   
   // Copy Cap from Main line to popup
   Sbr_INO_tConvoy_SL.rgtCap[Sbr_IN_dCapIndex].dColor := Sbr_INO_tConvoyCap_ZC.rgtCap[0].dColor;
   Sbr_INO_tConvoy_SL.rgtCap[Sbr_IN_dCapIndex].dConvTotLength_cmm := Sbr_INO_tConvoyCap_ZC.rgtCap[0].dConvTotLength_cmm;
   Sbr_INO_tConvoy_SL.rgtCap[Sbr_IN_dCapIndex].dFormat := Sbr_INO_tConvoyCap_ZC.rgtCap[0].dFormat;
   Sbr_INO_tConvoy_SL.rgtCap[Sbr_IN_dCapIndex].dGap_cmm := Sbr_INO_tConvoyCap_ZC.rgtCap[0].dGap_cmm;
   Sbr_INO_tConvoy_SL.rgtCap[Sbr_IN_dCapIndex].dID := Sbr_INO_tConvoyCap_ZC.rgtCap[0].dID;
   Sbr_INO_tConvoy_SL.rgtCap[Sbr_IN_dCapIndex].dIndex := Sbr_INO_tConvoyCap_ZC.rgtCap[0].dIndex;
   Sbr_INO_tConvoy_SL.rgtCap[Sbr_IN_dCapIndex].dLength_cmm := Sbr_INO_tConvoyCap_ZC.rgtCap[0].dLength_cmm;
   Sbr_INO_tConvoy_SL.rgtCap[Sbr_IN_dCapIndex].dMaxCapInConv := Sbr_INO_tConvoyCap_ZC.rgtCap[0].dMaxCapInConv;
   Sbr_INO_tConvoy_SL.rgtCap[Sbr_IN_dCapIndex].dNumLites := Sbr_INO_tConvoyCap_ZC.rgtCap[0].dNumLites;
   Sbr_INO_tConvoy_SL.rgtCap[Sbr_IN_dCapIndex].dProductionID := Sbr_INO_tConvoyCap_ZC.rgtCap[0].dProductionID;
   Sbr_INO_tConvoy_SL.rgtCap[Sbr_IN_dCapIndex].dReqGapForConv_cmm := Sbr_INO_tConvoyCap_ZC.rgtCap[0].dReqGapForConv_cmm;
   Sbr_INO_tConvoy_SL.rgtCap[Sbr_IN_dCapIndex].dStackerModality := Sbr_INO_tConvoyCap_ZC.rgtCap[0].dStackerModality;
   Sbr_INO_tConvoy_SL.rgtCap[Sbr_IN_dCapIndex].dStackerMode := Sbr_INO_tConvoyCap_ZC.rgtCap[0].dStackerMode;
   Sbr_INO_tConvoy_SL.rgtCap[Sbr_IN_dCapIndex].dThickness_cmm := Sbr_INO_tConvoyCap_ZC.rgtCap[0].dThickness_cmm;
   Sbr_INO_tConvoy_SL.rgtCap[Sbr_IN_dCapIndex].dWidth_cmm := Sbr_INO_tConvoyCap_ZC.rgtCap[0].dWidth_cmm;
   Sbr_INO_tConvoy_SL.rgtCap[Sbr_IN_dCapIndex].rgxDone := Sbr_INO_tConvoyCap_ZC.rgtCap[0].rgxDone;
   Sbr_INO_tConvoy_SL.rgtCap[Sbr_IN_dCapIndex].rgxRequest := Sbr_INO_tConvoyCap_ZC.rgtCap[0].rgxRequest;
   FOR TMP_dLite := 0 TO CONST_tPlant.dNumLitesMaxCap - 1 DO
   	Sbr_INO_tConvoy_SL.rgtCap[Sbr_IN_dCapIndex].rgtLite[TMP_dLite].dBarycenter_cmm := Sbr_INO_tConvoyCap_ZC.rgtCap[0].rgtLite[TMP_dLite].dBarycenter_cmm;
   	Sbr_INO_tConvoy_SL.rgtCap[Sbr_IN_dCapIndex].rgtLite[TMP_dLite].dCulletCause := Sbr_INO_tConvoyCap_ZC.rgtCap[0].rgtLite[TMP_dLite].dCulletCause;
   	Sbr_INO_tConvoy_SL.rgtCap[Sbr_IN_dCapIndex].rgtLite[TMP_dLite].dID := Sbr_INO_tConvoyCap_ZC.rgtCap[0].rgtLite[TMP_dLite].dID;
   	Sbr_INO_tConvoy_SL.rgtCap[Sbr_IN_dCapIndex].rgtLite[TMP_dLite].dProductionID := Sbr_INO_tConvoyCap_ZC.rgtCap[0].rgtLite[TMP_dLite].dProductionID;
   	Sbr_INO_tConvoy_SL.rgtCap[Sbr_IN_dCapIndex].rgtLite[TMP_dLite].dWidth_cmm := Sbr_INO_tConvoyCap_ZC.rgtCap[0].rgtLite[TMP_dLite].dWidth_cmm;
   	Sbr_INO_tConvoy_SL.rgtCap[Sbr_IN_dCapIndex].rgtLite[TMP_dLite].rgxDone := Sbr_INO_tConvoyCap_ZC.rgtCap[0].rgtLite[TMP_dLite].rgxDone;
   	Sbr_INO_tConvoy_SL.rgtCap[Sbr_IN_dCapIndex].rgtLite[TMP_dLite].rgxRequest := Sbr_INO_tConvoyCap_ZC.rgtCap[0].rgtLite[TMP_dLite].rgxRequest;
   	COP(Sbr_INO_tConvoyCap_ZC.rgtCap[0].rgtLite[TMP_dLite].tDestination,Sbr_INO_tConvoy_SL.rgtCap[Sbr_IN_dCapIndex].rgtLite[TMP_dLite].tDestination,1);
   	COP(Sbr_INO_tConvoyCap_ZC.rgtCap[0].rgtLite[TMP_dLite].tFlag,Sbr_INO_tConvoy_SL.rgtCap[Sbr_IN_dCapIndex].rgtLite[TMP_dLite].tFlag,1);
   END_FOR;
   Sbr_INO_tConvoy_SL.dLength_cmm := Sbr_INO_tConvoyCap_ZC.dLength_cmm;
   Sbr_INO_tConvoy_SL.dTotalCaps := Sbr_INO_tConvoyCap_ZC.dTotalCaps;
   Sbr_INO_tConvoy_SL.dGapCaps_cmm := Sbr_INO_tConvoyCap_ZC.dGapCaps_cmm;
   Sbr_INO_tConvoy_SL.dCapIndex := Sbr_INO_tConvoyCap_ZC.dCapIndex;
   Sbr_INO_tConvoy_SL.dNextCapIndex := Sbr_INO_tConvoyCap_ZC.dNextCapIndex;
   Sbr_IN_dCapIndex := Sbr_IN_dCapIndex + 1;
   
   // Call recursively to next cap
   IF Sbr_INO_tConvoyCap_ZC.dNextCapIndex > 0 AND Sbr_IN_dCapIndex < CONST_tPlant.dNumCapsMaxConvoy THEN
   	JSR(sbrConvDataLineToSL,3,Z300_BufferPlate.rgtPlate[Sbr_INO_tConvoyCap_ZC.dNextCapIndex].tData,Sbr_INO_tConvoy_SL,Sbr_IN_dCapIndex,Z300_BufferPlate.rgtPlate[Sbr_INO_tConvoyCap_ZC.dNextCapIndex].tData,Sbr_INO_tConvoy_SL);
   END_IF;
   
   //Output
   RET(Sbr_INO_tConvoyCap_ZC,Sbr_INO_tConvoy_SL);
   
END_ROUTINE

ROUTINE sbrConvDataSLToLine   (* structured text *)
   
   //Input
   SBR(Sbr_INO_tConvoyCap_ZC,Sbr_INO_tConvoy_SL,Sbr_IN_dCapIndex,Sbr_IN_ReentryPosition,Sbr_IN_ReentryPosition_min,Sbr_IN_ReentryPosition_max);
   
   COP(AUX_tConvoyCap_ZC_NULL,Sbr_INO_tConvoyCap_ZC,1);
   
   // Copy Cap from popup to main line
   Sbr_INO_tConvoyCap_ZC.rgtCap[0].dColor := Sbr_INO_tConvoy_SL.rgtCap[Sbr_IN_dCapIndex].dColor;
   Sbr_INO_tConvoyCap_ZC.rgtCap[0].dConvTotLength_cmm := Sbr_INO_tConvoy_SL.rgtCap[Sbr_IN_dCapIndex].dConvTotLength_cmm;
   Sbr_INO_tConvoyCap_ZC.rgtCap[0].dFormat := Sbr_INO_tConvoy_SL.rgtCap[Sbr_IN_dCapIndex].dFormat;
   Sbr_INO_tConvoyCap_ZC.rgtCap[0].dGap_cmm := Sbr_INO_tConvoy_SL.rgtCap[Sbr_IN_dCapIndex].dGap_cmm;
   Sbr_INO_tConvoyCap_ZC.rgtCap[0].dID := Sbr_INO_tConvoy_SL.rgtCap[Sbr_IN_dCapIndex].dID;
   Sbr_INO_tConvoyCap_ZC.rgtCap[0].dIndex := Sbr_INO_tConvoy_SL.rgtCap[Sbr_IN_dCapIndex].dIndex;
   Sbr_INO_tConvoyCap_ZC.rgtCap[0].dLength_cmm := Sbr_INO_tConvoy_SL.rgtCap[Sbr_IN_dCapIndex].dLength_cmm;
   Sbr_INO_tConvoyCap_ZC.rgtCap[0].dMaxCapInConv := Sbr_INO_tConvoy_SL.rgtCap[Sbr_IN_dCapIndex].dMaxCapInConv;
   Sbr_INO_tConvoyCap_ZC.rgtCap[0].dNumLites := Sbr_INO_tConvoy_SL.rgtCap[Sbr_IN_dCapIndex].dNumLites;
   Sbr_INO_tConvoyCap_ZC.rgtCap[0].dProductionID := Sbr_INO_tConvoy_SL.rgtCap[Sbr_IN_dCapIndex].dProductionID;
   Sbr_INO_tConvoyCap_ZC.rgtCap[0].dReqGapForConv_cmm := Sbr_INO_tConvoy_SL.rgtCap[Sbr_IN_dCapIndex].dReqGapForConv_cmm;
   Sbr_INO_tConvoyCap_ZC.rgtCap[0].dStackerModality := Sbr_INO_tConvoy_SL.rgtCap[Sbr_IN_dCapIndex].dStackerModality;
   Sbr_INO_tConvoyCap_ZC.rgtCap[0].dStackerMode := Sbr_INO_tConvoy_SL.rgtCap[Sbr_IN_dCapIndex].dStackerMode;
   Sbr_INO_tConvoyCap_ZC.rgtCap[0].dThickness_cmm := Sbr_INO_tConvoy_SL.rgtCap[Sbr_IN_dCapIndex].dThickness_cmm;
   Sbr_INO_tConvoyCap_ZC.rgtCap[0].dWidth_cmm := Sbr_INO_tConvoy_SL.rgtCap[Sbr_IN_dCapIndex].dWidth_cmm;
   Sbr_INO_tConvoyCap_ZC.rgtCap[0].rgxDone := Sbr_INO_tConvoy_SL.rgtCap[Sbr_IN_dCapIndex].rgxDone;
   Sbr_INO_tConvoyCap_ZC.rgtCap[0].rgxRequest := Sbr_INO_tConvoy_SL.rgtCap[Sbr_IN_dCapIndex].rgxRequest;
   FOR TMP_dLite := 0 TO CONST_tPlant.dNumLitesMaxCap - 1 DO
   	Sbr_INO_tConvoyCap_ZC.rgtCap[0].rgtLite[TMP_dLite].dBarycenter_cmm := Sbr_INO_tConvoy_SL.rgtCap[Sbr_IN_dCapIndex].rgtLite[TMP_dLite].dBarycenter_cmm;
   	Sbr_INO_tConvoyCap_ZC.rgtCap[0].rgtLite[TMP_dLite].dCulletCause := Sbr_INO_tConvoy_SL.rgtCap[Sbr_IN_dCapIndex].rgtLite[TMP_dLite].dCulletCause;
   	Sbr_INO_tConvoyCap_ZC.rgtCap[0].rgtLite[TMP_dLite].dID := Sbr_INO_tConvoy_SL.rgtCap[Sbr_IN_dCapIndex].rgtLite[TMP_dLite].dID;
   	Sbr_INO_tConvoyCap_ZC.rgtCap[0].rgtLite[TMP_dLite].dProductionID := Sbr_INO_tConvoy_SL.rgtCap[Sbr_IN_dCapIndex].rgtLite[TMP_dLite].dProductionID;
   	Sbr_INO_tConvoyCap_ZC.rgtCap[0].rgtLite[TMP_dLite].dWidth_cmm := Sbr_INO_tConvoy_SL.rgtCap[Sbr_IN_dCapIndex].rgtLite[TMP_dLite].dWidth_cmm;
   	Sbr_INO_tConvoyCap_ZC.rgtCap[0].rgtLite[TMP_dLite].rgxDone := Sbr_INO_tConvoy_SL.rgtCap[Sbr_IN_dCapIndex].rgtLite[TMP_dLite].rgxDone;
   	Sbr_INO_tConvoyCap_ZC.rgtCap[0].rgtLite[TMP_dLite].rgxRequest := Sbr_INO_tConvoy_SL.rgtCap[Sbr_IN_dCapIndex].rgtLite[TMP_dLite].rgxRequest;
   	COP(Sbr_INO_tConvoy_SL.rgtCap[Sbr_IN_dCapIndex].rgtLite[TMP_dLite].tDestination,Sbr_INO_tConvoyCap_ZC.rgtCap[0].rgtLite[TMP_dLite].tDestination,1);
   	COP(Sbr_INO_tConvoy_SL.rgtCap[Sbr_IN_dCapIndex].rgtLite[TMP_dLite].tFlag,Sbr_INO_tConvoyCap_ZC.rgtCap[0].rgtLite[TMP_dLite].tFlag,1);
   END_FOR;
   Sbr_INO_tConvoyCap_ZC.dLength_cmm := Sbr_INO_tConvoy_SL.dLength_cmm;
   Sbr_INO_tConvoyCap_ZC.dTotalCaps := Sbr_INO_tConvoy_SL.dTotalCaps;
   Sbr_INO_tConvoyCap_ZC.dGapCaps_cmm := Sbr_INO_tConvoy_SL.dGapCaps_cmm;
   Sbr_INO_tConvoyCap_ZC.dCapIndex := Sbr_INO_tConvoy_SL.dCapIndex;
   Sbr_INO_tConvoyCap_ZC.dNextCapIndex := 0;
   /////
   Sbr_IN_ReentryPosition := Sbr_IN_ReentryPosition - (Sbr_INO_tConvoy_SL.rgtCap[Sbr_IN_dCapIndex].dLength_cmm / 2);
   IF Sbr_IN_ReentryPosition < Sbr_IN_ReentryPosition_min THEN
   	Sbr_IN_ReentryPosition := Sbr_IN_ReentryPosition_min;
   END_IF;
   IF Sbr_IN_ReentryPosition > Sbr_IN_ReentryPosition_max THEN
   	Sbr_IN_ReentryPosition := Sbr_IN_ReentryPosition_max;
   END_IF;
   /////
   GP_TrackingAddCap(GP_TrackingAddCap,Z300_BufferPlate,Sbr_INO_tConvoyCap_ZC,Sbr_IN_ReentryPosition,0,-1,Z300_LineTracking,Z300_dEndTrackingPosition);
   TMP_rgdIndexC[Sbr_IN_dCapIndex] := GP_TrackingAddCap.OUT_dIndexInsertion;
   Sbr_IN_dCapIndex := Sbr_IN_dCapIndex + 1;
   
   // Call recursively to next cap
   IF Sbr_INO_tConvoy_SL.rgtCap[Sbr_IN_dCapIndex].dID > 0 AND Sbr_IN_dCapIndex < Sbr_INO_tConvoy_SL.dTotalCaps AND Sbr_IN_dCapIndex < CONST_tPlant.dNumCapsMaxConvoy THEN
   	IF Sbr_INO_tConvoy_SL.rgtCap[Sbr_IN_dCapIndex - 1].dReqGapForConv_cmm < CONST_tAux.dM302SpeedUpMinGapInConvoy_cmm THEN
   		Sbr_INO_tConvoy_SL.rgtCap[Sbr_IN_dCapIndex - 1].dReqGapForConv_cmm := CONST_tAux.dM302SpeedUpMinGapInConvoy_cmm;
   	END_IF;
   	Sbr_IN_ReentryPosition := Sbr_IN_ReentryPosition - Sbr_INO_tConvoy_SL.rgtCap[Sbr_IN_dCapIndex - 1].dLength_cmm - Sbr_INO_tConvoy_SL.rgtCap[Sbr_IN_dCapIndex - 1].dReqGapForConv_cmm;
   	JSR(sbrConvDataSLToLine,6,Sbr_INO_tConvoyCap_ZC,Sbr_INO_tConvoy_SL,Sbr_IN_dCapIndex,Sbr_IN_ReentryPosition,Sbr_IN_ReentryPosition_min,Sbr_IN_ReentryPosition_max);
   END_IF;
   
   //Output
   RET(Sbr_INO_tConvoyCap_ZC,Sbr_INO_tConvoy_SL);
   
END_ROUTINE

ROUTINE sbrForceData   (* structured text *)
   
   // only fortest
   //COP(AUX_tConvoyCapTest,Z200_SnapDataEth[0],1);
   //COP(AUX_tJumboTest,Z200_SnapDataEth[0],1);
   //////
   
   IF Z200_SnapDataEth[0].dLength_cmm <= 125000 THEN
   	Z200_SnapDataEth[0].rgtCap[0].dFormat := 2;
   	Z200_SnapDataEth[0].rgtCap[0].dStackerMode := 0;
   	Z200_SnapDataEth[0].rgtCap[0].dStackerModality := 10;
   END_IF;
   
   IF Z200_SnapDataEth[0].dLength_cmm <= 125000 AND Z200_SnapDataEth[0].rgtCap[0].rgtLite[0].dWidth_cmm = 140000 THEN
   	Z200_SnapDataEth[0].rgtCap[0].dFormat := 2;
   	Z200_SnapDataEth[0].rgtCap[0].dStackerMode := 0;
   	Z200_SnapDataEth[0].rgtCap[0].dStackerModality := 11;
   END_IF;
   
   IF Z200_SnapDataEth[0].dLength_cmm >= 600000 THEN
   	Z200_SnapDataEth[0].rgtCap[0].dFormat := 1;
   END_IF;
   
END_ROUTINE

ROUTINE sbrGetDataFromConvoy   (* structured text *)
   
   SBR(Sbr_IN_dIndexHead);
   
   Sbr_OUT_dTotalCaps := Z300_BufferPlate.rgtPlate[Sbr_IN_dIndexHead].tData.dTotalCaps;
   //initialize convoy data
   FOR TMP_dIndC := 0 TO 3 DO
   	Sbr_OUT_rgdConvoyLengths[TMP_dIndC] := 0;
   	IF TMP_dIndC < 3 THEN
   		Sbr_OUT_rgdConvoyGaps[TMP_dIndC] := 0;
   	END_IF;
   END_FOR;
   
   IF Sbr_OUT_dTotalCaps > 1 THEN
   	FOR TMP_dIndC := 0 TO Sbr_OUT_dTotalCaps - 1 DO
   		IF TMP_dIndC < 4 THEN
   			Sbr_OUT_rgdConvoyLengths[TMP_dIndC] := Z300_BufferPlate.rgtPlate[Sbr_IN_dIndexHead].tData.rgtCap[0].dLength_cmm;
   		END_IF;
   		IF ((TMP_dIndC < 3) AND (TMP_dIndC < (Sbr_OUT_dTotalCaps - 1))) THEN
   			Sbr_OUT_rgdConvoyGaps[TMP_dIndC] := Z300_BufferPlate.rgtPlate[Sbr_IN_dIndexHead].tData.rgtCap[0].dReqGapForConv_cmm;
   		END_IF;
   	END_FOR;
   END_IF;
   
   RET(Sbr_OUT_dTotalCaps,Sbr_OUT_rgdConvoyLengths,Sbr_OUT_rgdConvoyGaps);
   
END_ROUTINE

ROUTINE sbrM302CompileSnapData   (* structured text *)
   
   Z200_SnapDataEth[0].dGapCaps_cmm := 0;
   Z200_SnapDataEth[0].rgtCap[0].dGap_cmm := 0;
   Z200_SnapDataEth[0].rgtCap[0].dReqGapForConv_cmm := 0;
   Z200_SnapDataEth[0].dLength_cmm := Z200_SnapDataEth[0].rgtCap[0].dLength_cmm;
   IF Z200_SnapDataEth[0].dTotalCaps < 2 THEN //if single cap
   	Z200_SnapDataEth[0].rgtCap[0].dConvTotLength_cmm := Z200_SnapDataEth[0].rgtCap[0].dLength_cmm;
   ELSE //if convoy
   	Z200_SnapDataEth[0].dCapIndex := Z200_SnapDataEth[0].rgtCap[0].dIndex;
   	IF Z200_SnapDataEth[0].dCapIndex < ( Z200_SnapDataEth[0].dTotalCaps - 1) THEN
   		Z200_SnapDataEth[0].rgtCap[0].dReqGapForConv_cmm := M302SpeedUp.AUX_dStandardGap_cmm;
   	ELSE
   		Z200_SnapDataEth[0].rgtCap[0].dReqGapForConv_cmm := 0;
   	END_IF;
   	Z200_SnapDataEth[0].dGapCaps_cmm := Z200_SnapDataEth[0].rgtCap[0].dReqGapForConv_cmm;
   END_IF;
   
END_ROUTINE

ROUTINE sbrM302ConvoyCompleted   (* structured text *)
   
   //Initialize
   
   FOR TMP_d := 0 TO 4 DO
   	TMP_rgdPnt[TMP_d] := M302SpeedUp.tSearchPlate.rgdTailPointer[TMP_d];
   END_FOR;
   
   TMP_dPointer := TMP_rgdPnt[0];
   
   /*
   //Convoy Lenght
   IF M301SpeedUp.AUX_dNumCapConvoy > 1 THEN
       FOR TMP_dIndex := 0 TO M301SpeedUp.AUX_dNumCapConvoy - 1 DO
           TMP_dPointer := TMP_rgdPnt[TMP_dIndex];
           TMP_d := Z300_BufferPlate.rgtPlate[TMP_dPointer].tData.rgtCap[0].dLength_cmm + Z300_BufferPlate.rgtPlate[TMP_dPointer].tData.dGapCaps_cmm + TMP_d;
       END_FOR;
   END_IF;
   
   //Put data
   FOR TMP_dIndex := 0 TO M301SpeedUp.AUX_dNumCapConvoy - 1 DO
       TMP_dPointer := TMP_rgdPnt[TMP_dIndex];
       Z300_BufferPlate.rgtPlate[TMP_dPointer].tData.dLength_cmm := TMP_d;
   	//Z300_BufferPlate.rgtPlate[TMP_dPointer].tData.dTotalCaps := M301SpeedUp.AUX_dNumCapConvoy;
   	//Z300_BufferPlate.rgtPlate[TMP_dPointer].tData.rgtCap[0].dIndex := (M301SpeedUp.AUX_dNumCapConvoy - 1) - TMP_dIndex;
   	IF TMP_dIndex > 0 THEN
   		Z300_BufferPlate.rgtPlate[TMP_dPointer].tData.dNextCapIndex := TMP_rgdPnt[TMP_dIndex - 1];
   	END_IF;
   END_FOR;
   */
   
   //Find last plate of convoy
   IF (Z300_BufferPlate.rgtPlate[TMP_dPointer].tData.dTotalCaps > 1) AND (Z300_BufferPlate.rgtPlate[TMP_dPointer].tData.dCapIndex = Z300_BufferPlate.rgtPlate[TMP_dPointer].tData.dTotalCaps - 1) THEN
   	TMP_d := 0;
   	TMP_dConvoySearchMax := Z300_BufferPlate.rgtPlate[TMP_dPointer].tData.dTotalCaps;
   	//Convoy Lenght Calculation
       FOR TMP_dIndex := 0 TO TMP_dConvoySearchMax - 1 DO
           TMP_dPointer := TMP_rgdPnt[TMP_dIndex];
   		//////////////// Update dGapCaps with dReqGapForConv
   		Z300_BufferPlate.rgtPlate[TMP_dPointer].tData.dGapCaps_cmm := Z300_BufferPlate.rgtPlate[TMP_dPointer].tData.rgtCap[0].dReqGapForConv_cmm;
   		////////////////
           TMP_d := Z300_BufferPlate.rgtPlate[TMP_dPointer].tData.rgtCap[0].dLength_cmm + Z300_BufferPlate.rgtPlate[TMP_dPointer].tData.dGapCaps_cmm + TMP_d;
       END_FOR;
   	//From last plate of convoy set length and cap index next
   	FOR TMP_dIndex := 0 TO TMP_dConvoySearchMax - 1 DO
           TMP_dPointer := TMP_rgdPnt[TMP_dIndex];
   		Z300_BufferPlate.rgtPlate[TMP_dPointer].tData.dLength_cmm := TMP_d;
   		Z300_BufferPlate.rgtPlate[TMP_dPointer].tData.rgtCap[0].dConvTotLength_cmm := TMP_d;
   		//Set the next index if not last cap of convoy
   		IF (TMP_dIndex > 0) AND (Z300_BufferPlate.rgtPlate[TMP_dPointer].tData.dCapIndex < Z300_BufferPlate.rgtPlate[TMP_dPointer].tData.dTotalCaps - 1) THEN
   			Z300_BufferPlate.rgtPlate[TMP_dPointer].tData.dNextCapIndex := TMP_rgdPnt[TMP_dIndex - 1];
   			Z300_BufferPlate.rgtPlate[TMP_dPointer].tTracking.dNextCapIndex := TMP_rgdPnt[TMP_dIndex - 1];
   		ELSE
   			Z300_BufferPlate.rgtPlate[TMP_dPointer].tData.dNextCapIndex := 0;
   			Z300_BufferPlate.rgtPlate[TMP_dPointer].tTracking.dNextCapIndex := 0;
   		END_IF;
   		IF (TMP_dIndex < 3) AND (Z300_BufferPlate.rgtPlate[TMP_dPointer].tData.dCapIndex > 0)  THEN
   			Z300_BufferPlate.rgtPlate[TMP_dPointer].tTracking.dPreviousCapIndex := TMP_rgdPnt[TMP_dIndex + 1];
   		ELSE
   			Z300_BufferPlate.rgtPlate[TMP_dPointer].tTracking.dPreviousCapIndex := 0;
   		END_IF;
   	END_FOR;
   END_IF;
   
END_ROUTINE

ROUTINE sbrM302SnapCulletMissSnap   (* structured text *)
   
   //Set to cullet next cap to be snapped
   FOR TMP_dIndex:=0 TO CONST_tPlant.dNumLitesMaxCap - 1 DO
   	IF Z200_SnapDataEth[1].rgtCap[0].rgtLite[TMP_dIndex].dID <> 0 THEN
   		Z200_SnapDataEth[1].rgtCap[0].rgtLite[TMP_dIndex].tDestination.rgxMain := CONST_rgdDestMask[24];
   		//Interrupt convoy
   		Z200_SnapDataEth[1].rgtCap[0].dReqGapForConv_cmm := 0;
   		Z200_SnapDataEth[1].rgtCap[0].dIndex := 0;
   		M302SpeedUp.ST_xLastPlateInConvoy := 0;
   	END_IF;
   END_FOR;
   
END_ROUTINE

ROUTINE sbrM302SnapCulletWrongData   (* structured text *)
   
   FOR TMP_dIndex:=0 TO CONST_tPlant.dNumLitesMaxCap - 1 DO
   	IF Z200_SnapDataEth[1].rgtCap[0].rgtLite[TMP_dIndex].dID <> 0 THEN
   		Z200_SnapDataEth[1].rgtCap[0].rgtLite[TMP_dIndex].tDestination.rgxMain:=CONST_rgdDestMask[24];
   	END_IF;
   END_FOR;
   
END_ROUTINE

ROUTINE sbrM302SnapCulletWrongDim   (* structured text *)
   
   FOR TMP_dIndex:=0 TO CONST_tPlant.dNumLitesMaxCap - 1 DO
   	IF Z200_SnapDataEth[1].rgtCap[0].rgtLite[TMP_dIndex].dID <> 0 THEN
   		Z200_SnapDataEth[1].rgtCap[0].dLength_cmm := M302SpeedUp.AUX_dDimensionCapCreation_cmm;
   		Z200_SnapDataEth[1].rgtCap[0].rgtLite[TMP_dIndex].tDestination.rgxMain := CONST_rgdDestMask[24];
   	END_IF;
   END_FOR;
END_ROUTINE

ROUTINE sbrM30xPositionTrimFrame   (* ladder *)
   // #####_AUTOMATIC_POSITIONING_#####
   0: NOP();
   1: [XIC(M30xTrimDeck[TMP_dIndex].OS_xStartPositioning) ,XIC(M30xTrimDeck[TMP_dIndex].OS_xUpdateTarget) ][XIO(M30xTrimDeck_HMR[TMP_dIndex].xOpeningOnCleaningEnabled) ,XIC(M30xTrimDeck_HMR[TMP_dIndex].xOpeningOnCleaningEnabled) XIO(Z301.OS_xCleaningAccepted) XIO(Z301.ST_xCleaningAccepted) ]MOV(M30xTrimDeck_HMR[TMP_dIndex].rgdTarget_cmm[0],M30xTrimDeck[TMP_dIndex].AUX_dReqTargetPos_cmm[0])MOV(M30xTrimDeck_HMR[TMP_dIndex].rgdTarget_cmm[1],M30xTrimDeck[TMP_dIndex].AUX_dReqTargetPos_cmm[1])ADD(M30xTrimDeck[TMP_dIndex].AUX_dReqTargetPos_cmm[0],M30xTrimDeck[TMP_dIndex].AUX_dOffset_cmm[0],M30xTrimDeck[TMP_dIndex].AUX_dFinalTarget_cmm[0])ADD(M30xTrimDeck[TMP_dIndex].AUX_dReqTargetPos_cmm[1],M30xTrimDeck[TMP_dIndex].AUX_dOffset_cmm[1],M30xTrimDeck[TMP_dIndex].AUX_dFinalTarget_cmm[1]);
   2: GP_PosWindow(GP_PosWindow,M30xTrimDeck[TMP_dIndex].AUX_dFinalTarget_cmm[0],M30xTrimDeck[TMP_dIndex].AUX_dActTransPosition_cmm[0],M30xTrimDeck[TMP_dIndex].CONF_dTolerance_cmm,0,M30xTrimDeck[TMP_dIndex].ST_xInPositionOpSide)GP_PosWindow(GP_PosWindow,M30xTrimDeck[TMP_dIndex].AUX_dFinalTarget_cmm[1],M30xTrimDeck[TMP_dIndex].AUX_dActTransPosition_cmm[1],M30xTrimDeck[TMP_dIndex].CONF_dTolerance_cmm,0,M30xTrimDeck[TMP_dIndex].ST_xInPositionOppOpSide);
   3: GP_PosWindow(GP_PosWindow,M30xTrimDeck[TMP_dIndex].AUX_dFinalTarget_cmm[0],M30xTrimDeck[TMP_dIndex].AUX_dActTransPosition_cmm[0],M30xTrimDeck[TMP_dIndex].CONF_dSlowDown_cmm,0,M30xTrimDeck[TMP_dIndex].ST_xInSlowDownOpSide)GP_PosWindow(GP_PosWindow,M30xTrimDeck[TMP_dIndex].AUX_dFinalTarget_cmm[1],M30xTrimDeck[TMP_dIndex].AUX_dActTransPosition_cmm[1],M30xTrimDeck[TMP_dIndex].CONF_dSlowDown_cmm,0,M30xTrimDeck[TMP_dIndex].ST_xInSlowDownOppOpSide);
   4: GP_PosWindow(GP_PosWindow,M30xTrimDeck[TMP_dIndex].AUX_dFinalTarget_cmm[0],M30xTrimDeck[TMP_dIndex].AUX_dActTransPosition_cmm[0],M30xTrimDeck[TMP_dIndex].CONF_dStopCam_cmm,0,M30xTrimDeck[TMP_dIndex].ST_xStopCamPositionOpSide)GP_PosWindow(GP_PosWindow,M30xTrimDeck[TMP_dIndex].AUX_dFinalTarget_cmm[1],M30xTrimDeck[TMP_dIndex].AUX_dActTransPosition_cmm[1],M30xTrimDeck[TMP_dIndex].CONF_dStopCam_cmm,0,M30xTrimDeck[TMP_dIndex].ST_xStopCamPositionOppOpSide);
   // #####_MANUAL_POSITIONING_#####
   5: NOP();
   6: GP_PosWindow(GP_PosWindow,M30xTrimDeck_HMW[TMP_dIndex].dPositionManCmdOpSide_cmm,M30xTrimDeck[TMP_dIndex].AUX_dActTransPosition_cmm[0],M30xTrimDeck[TMP_dIndex].CONF_dSlowDown_cmm,0,M30xTrimDeck[TMP_dIndex].ST_xInSlowDownManualOpSide)GP_PosWindow(GP_PosWindow,M30xTrimDeck_HMW[TMP_dIndex].dPositionManCmdOpSide_cmm,M30xTrimDeck[TMP_dIndex].AUX_dActTransPosition_cmm[1],M30xTrimDeck[TMP_dIndex].CONF_dSlowDown_cmm,0,M30xTrimDeck[TMP_dIndex].ST_xInSlowDownManualOppOpSide);
   7: GP_PosWindow(GP_PosWindow,M30xTrimDeck[TMP_dIndex].AUX_dFinalTarget_cmm[0],M30xTrimDeck[TMP_dIndex].AUX_dActTransPosition_cmm[0],M30xTrimDeck[TMP_dIndex].CONF_dStopCam_cmm,0,M30xTrimDeck[TMP_dIndex].ST_xStopCamManualPositionOpSide)GP_PosWindow(GP_PosWindow,M30xTrimDeck[TMP_dIndex].AUX_dFinalTarget_cmm[1],M30xTrimDeck[TMP_dIndex].AUX_dActTransPosition_cmm[1],M30xTrimDeck[TMP_dIndex].CONF_dStopCam_cmm,0,M30xTrimDeck[TMP_dIndex].ST_xStopCamManualPositionOppOpSide);
   8: XIC(M30xTrimDeck_HMW[TMP_dIndex].rgxMan.x0)MOV(M30xTrimDeck[TMP_dIndex].CONF_dTrimDeckMinPos_cmm[0],TMP_dManualTargetPos);
   9: XIC(M30xTrimDeck_HMW[TMP_dIndex].rgxMan.x1)MOV(M30xTrimDeck[TMP_dIndex].CONF_dTrimDeckMaxPos_cmm[0],TMP_dManualTargetPos);
   10: XIC(M30xTrimDeck_HMW[TMP_dIndex].rgxMan.x4)MOV(M30xTrimDeck[TMP_dIndex].CONF_dTrimDeckMinPos_cmm[1],TMP_dManualTargetPos);
   11: XIC(M30xTrimDeck_HMW[TMP_dIndex].rgxMan.x5)MOV(M30xTrimDeck[TMP_dIndex].CONF_dTrimDeckMaxPos_cmm[1],TMP_dManualTargetPos);
   12: GP_PosWindow(GP_PosWindow,TMP_dManualTargetPos,M30xTrimDeck[TMP_dIndex].AUX_dActTransPosition_cmm[0],M30xTrimDeck[TMP_dIndex].CONF_dSlowDown_cmm,0,M30xTrimDeck[TMP_dIndex].ST_xInSlowDownManualOpSide)GP_PosWindow(GP_PosWindow,TMP_dManualTargetPos,M30xTrimDeck[TMP_dIndex].AUX_dActTransPosition_cmm[1],M30xTrimDeck[TMP_dIndex].CONF_dSlowDown_cmm,0,M30xTrimDeck[TMP_dIndex].ST_xInSlowDownManualOppOpSide);
   13: GP_PosWindow(GP_PosWindow,TMP_dManualTargetPos,M30xTrimDeck[TMP_dIndex].AUX_dActTransPosition_cmm[0],M30xTrimDeck[TMP_dIndex].CONF_dStopCam_cmm,0,M30xTrimDeck[TMP_dIndex].ST_xStopCamManualPositionOpSide)GP_PosWindow(GP_PosWindow,TMP_dManualTargetPos,M30xTrimDeck[TMP_dIndex].AUX_dActTransPosition_cmm[1],M30xTrimDeck[TMP_dIndex].CONF_dStopCam_cmm,0,M30xTrimDeck[TMP_dIndex].ST_xStopCamManualPositionOppOpSide);
END_ROUTINE

ROUTINE sbrM30xTrimDeckFramePositioning   (* ladder *)
   0: NOP();
   1: [NEQ(M30xTrimDeck_DATA[TMP_dIndex].rgtCap[0].dMaxWidth_cmm,M30xTrimDeck_DATA[TMP_dIndex].rgtCap[0].dMinWidth_cmm) [OTE(M30xTrimDeck[TMP_dIndex].ST_xDoubleSizeProduction) ,CPT(M303_dHalfWidthDifference,(M30xTrimDeck_DATA[TMP_dIndex].rgtCap[0].dMaxWidth_cmm - M30xTrimDeck_DATA[TMP_dIndex].rgtCap[0].dMinWidth_cmm) / 2) ] ,GEQ(M30xTrimDeck_DATA[TMP_dIndex].rgtCap[0].dLength_cmm,CONST_tPlant.rgdLiteLimits_cmm[4]) OTE(M30xTrimDeck[TMP_dIndex].ST_xJumboInProgress) ,[GRT(M30xTrimDeck_DATA[TMP_dIndex].dTotalCaps,1) ,GRT(M30xTrimDeck_DATA[TMP_dIndex].rgtCap[0].dIndex,0) ] OTE(M30xTrimDeck[TMP_dIndex].ST_xConvoyInProgress) ,EQU(M30xTrimDeck_DATA[TMP_dIndex].rgtCap[0].dIndex,0) OTE(M30xTrimDeck[TMP_dIndex].ST_xFirstCapInConv) ,[EQU(M30xTrimDeck_DATA[TMP_dIndex].rgtCap[0].rgtLite[0].tDestination.rgxMain,CONST_rgdDestMask[29]) ,EQU(M30xTrimDeck_DATA[TMP_dIndex].rgtCap[0].rgtLite[0].tDestination.rgxMain,CONST_rgdDestMask[30]) ,EQU(M30xTrimDeck_DATA[TMP_dIndex].rgtCap[0].rgtLite[0].tDestination.rgxMain,CONST_rgdDestMask[31]) ] OTE(M30xTrimDeck[TMP_dIndex].ST_xQualityInProgress) ,LEQ(M30xTrimDeck_DATA[TMP_dIndex].rgtCap[0].dNumLites,1) EQU(M30xTrimDeck_DATA[TMP_dIndex].rgtCap[0].rgtLite[0].tDestination.rgxMain,CONST_rgdDestMask[24]) OTE(M30xTrimDeck[TMP_dIndex].ST_xCulletInProgress) ,XIC(M30xTrimDeck[TMP_dIndex].ST_xDoubleSizeProduction) [CMP(M30xTrimDeck_DATA[TMP_dIndex].rgtCap[0].dWidth_cmm <= (M30xTrimDeck_DATA[TMP_dIndex].rgtCap[0].dMaxWidth_cmm + M30xTrimDeck_DATA[TMP_dIndex].rgtCap[0].dMinWidth_cmm) / 2) OTE(M30xTrimDeck[TMP_dIndex].ST_xShortestInProgress) ,CMP(M30xTrimDeck_DATA[TMP_dIndex].rgtCap[0].dWidth_cmm > (M30xTrimDeck_DATA[TMP_dIndex].rgtCap[0].dMaxWidth_cmm + M30xTrimDeck_DATA[TMP_dIndex].rgtCap[0].dMinWidth_cmm) / 2) OTE(M30xTrimDeck[TMP_dIndex].ST_xBiggestInProgress) ] ];
   2: [XIO(M30xTrimDeck[TMP_dIndex].ST_xConvoyInProgress) ,XIC(M30xTrimDeck[TMP_dIndex].ST_xFirstCapInConv) ][[XIC(M30xTrimDeck_DATA[TMP_dIndex].rgtCap[0].tFlag.xTrim3OpSide) ,XIC(M30xTrimDeck_DATA[TMP_dIndex].rgtCap[0].tFlag.xTrim2OpSide) ,XIC(M30xTrimDeck_DATA[TMP_dIndex].rgtCap[0].tFlag.xTrim1OpSide) ] OTE(M30xTrimDeck[TMP_dIndex].ST_xTrimDeckInWorkOpSide) ,[XIC(M30xTrimDeck_DATA[TMP_dIndex].rgtCap[0].tFlag.xTrim1OppOpSide) ,XIC(M30xTrimDeck_DATA[TMP_dIndex].rgtCap[0].tFlag.xTrim2OppOpSide) ,XIC(M30xTrimDeck_DATA[TMP_dIndex].rgtCap[0].tFlag.xTrim3OppOpSide) ] OTE(M30xTrimDeck[TMP_dIndex].ST_xTrimDeckInWorkOppOpSide) ];
   // Check wander limits
   3: XIC(M30xTrimDeck_HMR[TMP_dIndex].xControlWanderEnabled)[MOV(M30xTrimDeck_DATA[TMP_dIndex].rgtCap[0].dCutWander_cmm,TMP_dWander) ,LES(M30xTrimDeck_DATA[TMP_dIndex].rgtCap[0].dCutWander_cmm,CONST_tPlant.rgdWanderLimits[0]) MOV(CONST_tPlant.rgdWanderLimits[0],TMP_dWander) ,GRT(M30xTrimDeck_DATA[TMP_dIndex].rgtCap[0].dCutWander_cmm,CONST_tPlant.rgdWanderLimits[1]) MOV(CONST_tPlant.rgdWanderLimits[1],TMP_dWander) ];
   // Calculate target position with machine in work
   4: [XIC(M30xTrimDeck[TMP_dIndex].OS_xStartMoveFromTracking) ,XIC(M30xTrimDeck[TMP_dIndex].OS_xStartMoveFromEth1) ,XIC(M30xTrimDeck[TMP_dIndex].ST_xReqStartMovement) ][XIC(M30xTrimDeck[TMP_dIndex].ST_xTrimDeckInWorkOpSide) ,XIC(M30xTrimDeck[TMP_dIndex].ST_xTrimDeckInWorkOppOpSide) ]OTE(TMP_x);
   5: XIC(TMP_x)[DIV(M30xTrimDeck[TMP_dIndex].CONF_dTrimDeckMinRange_cmm,2,M30xTrimDeck[TMP_dIndex].AUX_dTarget_cmm[0]) ,GRT(M30xTrimDeck_DATA[TMP_dIndex].rgtCap[0].dWidth_cmm,M30xTrimDeck[TMP_dIndex].CONF_dTrimDeckMinRange_cmm) [DIV(M30xTrimDeck_DATA[TMP_dIndex].rgtCap[0].dWidth_cmm,2,M30xTrimDeck[TMP_dIndex].AUX_dTarget_cmm[0]) GRT(M30xTrimDeck_DATA[TMP_dIndex].rgtCap[0].dMinWidth_cmm,0) DIV(M30xTrimDeck_DATA[TMP_dIndex].rgtCap[0].dMinWidth_cmm,2,M30xTrimDeck[TMP_dIndex].AUX_dTarget_cmm[0]) ,[XIO(M30xTrimDeck[TMP_dIndex].ST_xDoubleSizeProduction) ,XIC(M30xTrimDeck_DATA[TMP_dIndex].rgtCap[0].tFlag.xOptSelvedgeSel) ] [XIO(M30xTrimDeck[TMP_dIndex].ST_xJumboInProgress) ,XIO(xAlwaysOFF) ] [XIC(M30xTrimDeck_DATA[TMP_dIndex].rgtCap[0].tFlag.xTrim2OpSide) ,XIC(M30xTrimDeck_DATA[TMP_dIndex].rgtCap[0].tFlag.xTrim3OpSide) ] XIC(xAlwaysOFF) ADD(M30xTrimDeck[TMP_dIndex].AUX_dTarget_cmm[0],M30xTrimDeck_DATA[TMP_dIndex].rgtCap[0].dDEdgeOpSide_cmm,M30xTrimDeck[TMP_dIndex].AUX_dTarget_cmm[0]) ] ,XIC(M30xTrimDeck_HMR[TMP_dIndex].xControlWanderEnabled) SUB(M30xTrimDeck[TMP_dIndex].AUX_dTarget_cmm[0],TMP_dWander,M30xTrimDeck[TMP_dIndex].AUX_dTarget_cmm[0]) ];
   6: XIC(TMP_x)[DIV(M30xTrimDeck[TMP_dIndex].CONF_dTrimDeckMinRange_cmm,2,M30xTrimDeck[TMP_dIndex].AUX_dTarget_cmm[1]) ,GRT(M30xTrimDeck_DATA[TMP_dIndex].rgtCap[0].dWidth_cmm,M30xTrimDeck[TMP_dIndex].CONF_dTrimDeckMinRange_cmm) [DIV(M30xTrimDeck_DATA[TMP_dIndex].rgtCap[0].dWidth_cmm,2,M30xTrimDeck[TMP_dIndex].AUX_dTarget_cmm[1]) GRT(M30xTrimDeck_DATA[TMP_dIndex].rgtCap[0].dMinWidth_cmm,0) DIV(M30xTrimDeck_DATA[TMP_dIndex].rgtCap[0].dMinWidth_cmm,2,M30xTrimDeck[TMP_dIndex].AUX_dTarget_cmm[1]) ,[XIO(M30xTrimDeck[TMP_dIndex].ST_xDoubleSizeProduction) ,XIC(M30xTrimDeck_DATA[TMP_dIndex].rgtCap[0].tFlag.xOptSelvedgeSel) ] [XIO(M30xTrimDeck[TMP_dIndex].ST_xJumboInProgress) ,XIO(xAlwaysOFF) ] [XIC(M30xTrimDeck_DATA[TMP_dIndex].rgtCap[0].tFlag.xTrim2OppOpSide) ,XIC(M30xTrimDeck_DATA[TMP_dIndex].rgtCap[0].tFlag.xTrim3OppOpSide) ] XIC(xAlwaysOFF) ADD(M30xTrimDeck[TMP_dIndex].AUX_dTarget_cmm[1],M30xTrimDeck_DATA[TMP_dIndex].rgtCap[0].dDEdgeOppOpSide_cmm,M30xTrimDeck[TMP_dIndex].AUX_dTarget_cmm[1]) ] ,XIC(M30xTrimDeck_HMR[TMP_dIndex].xControlWanderEnabled) ADD(M30xTrimDeck[TMP_dIndex].AUX_dTarget_cmm[1],TMP_dWander,M30xTrimDeck[TMP_dIndex].AUX_dTarget_cmm[1]) ];
   7: [XIC(TMP_x) MOV(M30xTrimDeck_DATA[TMP_dIndex].rgtCap[0].dWidth_cmm,M30xTrimDeck_HMR[TMP_dIndex].dNetWidthInProgress_cmm) MOV(M30xTrimDeck_DATA[TMP_dIndex].rgtCap[0].dGrossWidth_cmm,M30xTrimDeck_HMR[TMP_dIndex].dGrossWidthInProgress_cmm) MOV(M30xTrimDeck_DATA[TMP_dIndex].rgtCap[0].dCutWander_cmm,M30xTrimDeck_HMR[TMP_dIndex].dCutWanderInProgress_cmm) ,XIO(TMP_x) MOV(0,M30xTrimDeck_HMR[TMP_dIndex].dNetWidthInProgress_cmm) MOV(0,M30xTrimDeck_HMR[TMP_dIndex].dGrossWidthInProgress_cmm) MOV(0,M30xTrimDeck_HMR[TMP_dIndex].dCutWanderInProgress_cmm) ];
   // Calculate target position with machine in rest
   8: XIC(M30xTrimDeck[TMP_dIndex].ST_xReqStartMovement)XIO(M30xTrimDeck[TMP_dIndex].ST_xTrimDeckInWorkOpSide)XIO(M30xTrimDeck[TMP_dIndex].ST_xTrimDeckInWorkOppOpSide)OTE(TMP_x);
   9: XIC(TMP_x)[XIC(xAlwaysOFF) XIC(M30xTrimDeck_HMR[TMP_dIndex].xControlWanderEnabled) SUB(M30xTrimDeck[TMP_dIndex].AUX_dTarget_cmm[0],M30xTrimDeck_HMR[TMP_dIndex].dCutWanderInProgress_cmm,M30xTrimDeck[TMP_dIndex].AUX_dTarget_cmm[0]) XIC(xAlwaysOFF) NEQ(M30xTrimDeck_HMR[TMP_dIndex].dCutWanderInProgress_cmm,TMP_dWander) CPT(M30xTrimDeck[TMP_dIndex].AUX_dTarget_cmm[0],M30xTrimDeck[TMP_dIndex].AUX_dTarget_cmm[0] + (M30xTrimDeck_HMR[TMP_dIndex].dCutWanderInProgress_cmm - TMP_dWander)) ,XIC(xAlwaysOFF) CMP(M30xTrimDeck_DATA[TMP_dIndex].rgtCap[0].dWidth_cmm > M30xTrimDeck_HMR[TMP_dIndex].dDistBetweenSides_cmm + ((M30xTrimDeck[TMP_dIndex].CONF_dTrimDeckWheelsDist_cmm[0] + M30xTrimDeck[TMP_dIndex].CONF_dTrimDeckWheelsDist_cmm[1])/2)) GRT(M30xTrimDeck_DATA[TMP_dIndex].rgtCap[0].dWidth_cmm,M30xTrimDeck[TMP_dIndex].CONF_dTrimDeckMinRange_cmm) [CPT(M30xTrimDeck[TMP_dIndex].AUX_dTarget_cmm[0],(M30xTrimDeck_DATA[TMP_dIndex].rgtCap[0].dWidth_cmm + (M30xTrimDeck[TMP_dIndex].CONF_dTrimDeckWheelsDist_cmm[0] + M30xTrimDeck[TMP_dIndex].CONF_dTrimDeckWheelsDist_cmm[1])/2)/2) ,XIC(M30xTrimDeck_HMR[TMP_dIndex].xControlWanderEnabled) SUB(M30xTrimDeck[TMP_dIndex].AUX_dTarget_cmm[0],TMP_dWander,M30xTrimDeck[TMP_dIndex].AUX_dTarget_cmm[0]) ] ];
   10: XIC(TMP_x)[XIC(xAlwaysOFF) XIC(M30xTrimDeck_HMR[TMP_dIndex].xControlWanderEnabled) ADD(M30xTrimDeck[TMP_dIndex].AUX_dTarget_cmm[1],M30xTrimDeck_HMR[TMP_dIndex].dCutWanderInProgress_cmm,M30xTrimDeck[TMP_dIndex].AUX_dTarget_cmm[1]) XIC(xAlwaysOFF) NEQ(M30xTrimDeck_HMR[TMP_dIndex].dCutWanderInProgress_cmm,TMP_dWander) CPT(M30xTrimDeck[TMP_dIndex].AUX_dTarget_cmm[1],M30xTrimDeck[TMP_dIndex].AUX_dTarget_cmm[1] - (M30xTrimDeck_HMR[TMP_dIndex].dCutWanderInProgress_cmm - TMP_dWander)) ,XIC(xAlwaysOFF) CMP(M30xTrimDeck_DATA[TMP_dIndex].rgtCap[0].dWidth_cmm > M30xTrimDeck_HMR[TMP_dIndex].dDistBetweenSides_cmm + ((M30xTrimDeck[TMP_dIndex].CONF_dTrimDeckWheelsDist_cmm[0] + M30xTrimDeck[TMP_dIndex].CONF_dTrimDeckWheelsDist_cmm[1])/2)) GRT(M30xTrimDeck_DATA[TMP_dIndex].rgtCap[0].dWidth_cmm,M30xTrimDeck[TMP_dIndex].CONF_dTrimDeckMinRange_cmm) [CPT(M30xTrimDeck[TMP_dIndex].AUX_dTarget_cmm[1],(M30xTrimDeck_DATA[TMP_dIndex].rgtCap[0].dWidth_cmm + (M30xTrimDeck[TMP_dIndex].CONF_dTrimDeckWheelsDist_cmm[0] + M30xTrimDeck[TMP_dIndex].CONF_dTrimDeckWheelsDist_cmm[1])/2)/2) ,XIC(M30xTrimDeck_HMR[TMP_dIndex].xControlWanderEnabled) ADD(M30xTrimDeck[TMP_dIndex].AUX_dTarget_cmm[1],TMP_dWander,M30xTrimDeck[TMP_dIndex].AUX_dTarget_cmm[1]) ] ];
   // Offset calculations
   11: XIC(M30xTrimDeck_HMR[TMP_dIndex].xControlWidthEnabled)XIC(M30xTrimDeck[TMP_dIndex].ST_xOutputEnable)[XIC(M30xTrimDeck[TMP_dIndex].INPUT_xSATrimDeckToExternal.0) ,XIC(M30xTrimDeck[TMP_dIndex].INPUT_xSATrimDeckToExternal.10) ]ONS(M30xTrimDeck[TMP_dIndex].OSR_xOpSideToExternal)XIO(M30xTrimDeck[TMP_dIndex].INPUT_xSQTrimDeckExternalStop.0)LES(M30xTrimDeck_HMR[TMP_dIndex].rgdPosition_cmm[0],M30xTrimDeck[TMP_dIndex].CONF_dTrimDeckMaxPos_cmm[0])LES(M30xTrimDeck_HMR[TMP_dIndex].dDistBetweenSides_cmm,M30xTrimDeck[TMP_dIndex].CONF_dTrimDeckMaxRange_cmm)ADD(M30xTrimDeck_HMR[TMP_dIndex].rgdOffsetEachSide_cmm[0],M30xTrimDeck_HMW[TMP_dIndex].dOffsetOpSide_cmm,M30xTrimDeck_HMR[TMP_dIndex].rgdOffsetEachSide_cmm[0]);
